// TIA Portal project "liftvezerles" (V17)
// Az Automatizálási Tanszék SIMATIC eszközei

(* hardware
DEVICE "S7-1200 station_1"  S7-1200 Station
   slot 0: "Rack_0"  S7-1200 Rack  Rack  V1.0
   slot 1: "S71214_sim"  CPU 1214C DC/DC/DC  6ES7 214-1AG40-0XB0  V4.0
   slot 3: "AQ 1x12BIT_1"  AQ1 signal board  6ES7 232-4HA30-0XB0  V1.0
DEVICE "KTP700.Basic"  KTP700 Basic PN
   slot 0: "KTP700.Basic"  KTP700 Basic PN  6AV2 123-2GB03-0AX0  17.0.0.0
   slot 1: "HMI_RT_1"  KTP700 Basic PN  6AV2 123-2GB03-0AX0  17.0.0.0
   slot 5: "KTP700.Basic.IE_CP_1"  PROFINET Interface  17.0.0.0
      slot 1: "PROFINET Interface_1"  PROFINET Interface
         slot 1: "Port_1"  Port
DEVICE "S7-1200 station_2"  S7-1200 Station
   slot 0: "Rack_0"  S7-1200 Rack  Rack  V1.0
   slot 1: "S7.1214_aut"  CPU 1214C DC/DC/DC  6ES7 214-1AG31-0XB0  V3.0
   slot 3: "AQ 1x12BIT_1"  AQ1 signal board  6ES7 232-4HA30-0XB0  V1.0
*)

// ===== PLC "S71214_sim"  CPU 1214C DC/DC/DC =====

VAR_GLOBAL   // PLC tag table "Default tag table"
   "System_Byte" AT %MB11 : Byte;
   "FirstScan" AT %M11.0 : Bool;
   "DiagStatusUpdate" AT %M11.1 : Bool;
   "AlwaysTRUE" AT %M11.2 : Bool;
   "AlwaysFALSE" AT %M11.3 : Bool;
   "Clock_Byte" AT %MB10 : Byte;
   "Clock_10Hz" AT %M10.0 : Bool;
   "Clock_5Hz" AT %M10.1 : Bool;
   "Clock_2.5Hz" AT %M10.2 : Bool;
   "Clock_2Hz" AT %M10.3 : Bool;
   "Clock_1.25Hz" AT %M10.4 : Bool;
   "Clock_1Hz" AT %M10.5 : Bool;
   "Clock_0.625Hz" AT %M10.6 : Bool;
   "Clock_0.5Hz" AT %M10.7 : Bool;
END_VAR

VAR_GLOBAL   // PLC tag table "Elevatorcontrol"
   "elevator1position" AT %MW28 : Int;
   "elevator2position" AT %MW26 : Int;
END_VAR

VAR_GLOBAL   // PLC tag table "IO"
   "door1closemotor" AT %M8.0 : Bool;
   "door2openmotor" AT %M8.1 : Bool;
   "door1opensens" AT %M8.2 : Bool;
   "door1closedsens" AT %M8.3 : Bool;
   "door2opensens" AT %M8.4 : Bool;
   "door2closedsens" AT %M8.5 : Bool;
   "door1openmotor" AT %M8.6 : Bool;
   "door2closemotor" AT %M8.7 : Bool;
   "elevator1upmotor" AT %M9.0 : Bool;
   "elevator1downmotor" AT %M9.1 : Bool;
   "elevator2upmotor" AT %M9.2 : Bool;
   "elevator2downmotor" AT %M9.3 : Bool;
   "proximity1ground" AT %M9.4 : Bool;
   "proximity11" AT %M9.5 : Bool;
   "proximity12" AT %M9.6 : Bool;
   "proximity13" AT %M9.7 : Bool;
   "proximity14" AT %M12.0 : Bool;
   "proximity15" AT %M12.1 : Bool;
   "proximity2ground" AT %M12.2 : Bool;
   "proximity21" AT %M12.3 : Bool;
   "proximity22" AT %M12.4 : Bool;
   "proximity23" AT %M12.5 : Bool;
   "proximity24" AT %M12.6 : Bool;
   "proximity25" AT %M12.7 : Bool;
END_VAR

VAR_GLOBAL   // PLC tag table "HMI_IO"
   "requpgnd" AT %M7.0 : Bool;
   "requp1" AT %M7.1 : Bool;
   "requp2" AT %M7.2 : Bool;
   "requp3" AT %M7.3 : Bool;
   "requp4" AT %M7.4 : Bool;
   "reqdown5" AT %M7.5 : Bool;
   "reqdown4" AT %M7.6 : Bool;
   "reqdown3" AT %M7.7 : Bool;
   "reqdown2" AT %M5.6 : Bool;
   "reqdown1" AT %M5.7 : Bool;
   "req10" AT %M4.2 : Bool;
   "req11" AT %M4.3 : Bool;
   "req12" AT %M4.4 : Bool;
   "req13" AT %M4.5 : Bool;
   "req14" AT %M4.6 : Bool;
   "req15" AT %M4.7 : Bool;
   "req20" AT %M5.0 : Bool;
   "req21" AT %M5.1 : Bool;
   "req22" AT %M5.2 : Bool;
   "req23" AT %M5.3 : Bool;
   "req24" AT %M5.4 : Bool;
   "req25" AT %M5.5 : Bool;
   "las2" AT %M6.1 : Bool;
   "las1" AT %M6.0 : Bool;
   "doorclosebutton1" AT %M6.2 : Bool;
   "doorclosebutton2" AT %M6.3 : Bool;
   "dooropenbutton1" AT %M6.4 : Bool;
   "dooropenbutton2" AT %M6.5 : Bool;
END_VAR

VAR_GLOBAL   // PLC tag table "IO_simulation_tags"
   "lastfloor1" AT %MW18 : Int;
   "lastfloor2" AT %MW20 : Int;
   "state1" AT %MW22 : Int;
   "state2" AT %MW24 : Int;
   "elevator1positionsim" AT %MW14 : Int;
   "elevator2positionsim" AT %MW16 : Int;
END_VAR

VAR_GLOBAL   // PLC tag table "HMI_display_tags"
   "activefloor" AT %MW40 : Int;
   "door1open" AT %M42.0 : Bool;
   "door2open" AT %M42.1 : Bool;
END_VAR

DATA_BLOCK "ControlBlock_DB"   // DB9
{ S7_Optimized_Access := 'TRUE' }
VERSION : 0.1
// stored: InstanceOfName ControlBlock
"ControlBlock"
BEGIN
END_DATA_BLOCK

// folder: System blocks/Program resources

DATA_BLOCK "door1closing"   // DB5
{ S7_Optimized_Access := 'TRUE' }
AUTHOR : Simatic
FAMILY : IEC
NAME : IEC_TMR
VERSION : 1.0
// stored: InstanceOfName IEC_TIMER
"IEC_TIMER"
BEGIN
END_DATA_BLOCK

DATA_BLOCK "door1opening"   // DB6
{ S7_Optimized_Access := 'TRUE' }
AUTHOR : Simatic
FAMILY : IEC
NAME : IEC_TMR
VERSION : 1.0
// stored: InstanceOfName IEC_TIMER
"IEC_TIMER"
BEGIN
END_DATA_BLOCK

DATA_BLOCK "door2closing"   // DB7
{ S7_Optimized_Access := 'TRUE' }
AUTHOR : Simatic
FAMILY : IEC
NAME : IEC_TMR
VERSION : 1.0
// stored: InstanceOfName IEC_TIMER
"IEC_TIMER"
BEGIN
END_DATA_BLOCK

DATA_BLOCK "door2opening"   // DB8
{ S7_Optimized_Access := 'TRUE' }
AUTHOR : Simatic
FAMILY : IEC
NAME : IEC_TMR
VERSION : 1.0
// stored: InstanceOfName IEC_TIMER
"IEC_TIMER"
BEGIN
END_DATA_BLOCK

DATA_BLOCK "starting_up2"   // DB10
{ S7_Optimized_Access := 'TRUE' }
AUTHOR : Simatic
FAMILY : IEC
NAME : IEC_TMR
VERSION : 1.0
// stored: InstanceOfName IEC_TIMER
"IEC_TIMER"
BEGIN
END_DATA_BLOCK

DATA_BLOCK "starting_down2"   // DB11
{ S7_Optimized_Access := 'TRUE' }
AUTHOR : Simatic
FAMILY : IEC
NAME : IEC_TMR
VERSION : 1.0
// stored: InstanceOfName IEC_TIMER
"IEC_TIMER"
BEGIN
END_DATA_BLOCK

DATA_BLOCK "goingup2"   // DB12
{ S7_Optimized_Access := 'TRUE' }
AUTHOR : Simatic
FAMILY : IEC
NAME : IEC_TMR
VERSION : 1.0
// stored: InstanceOfName IEC_TIMER
"IEC_TIMER"
BEGIN
END_DATA_BLOCK

DATA_BLOCK "goingdown2"   // DB13
{ S7_Optimized_Access := 'TRUE' }
AUTHOR : Simatic
FAMILY : IEC
NAME : IEC_TMR
VERSION : 1.0
// stored: InstanceOfName IEC_TIMER
"IEC_TIMER"
BEGIN
END_DATA_BLOCK

DATA_BLOCK "starting_up1"   // DB20
{ S7_Optimized_Access := 'TRUE' }
AUTHOR : Simatic
FAMILY : IEC
NAME : IEC_TMR
VERSION : 1.0
// stored: InstanceOfName IEC_TIMER
"IEC_TIMER"
BEGIN
END_DATA_BLOCK

DATA_BLOCK "starting_down1"   // DB21
{ S7_Optimized_Access := 'TRUE' }
AUTHOR : Simatic
FAMILY : IEC
NAME : IEC_TMR
VERSION : 1.0
// stored: InstanceOfName IEC_TIMER
"IEC_TIMER"
BEGIN
END_DATA_BLOCK

DATA_BLOCK "goingup1"   // DB22
{ S7_Optimized_Access := 'TRUE' }
AUTHOR : Simatic
FAMILY : IEC
NAME : IEC_TMR
VERSION : 1.0
// stored: InstanceOfName IEC_TIMER
"IEC_TIMER"
BEGIN
END_DATA_BLOCK

DATA_BLOCK "goingdown1"   // DB23
{ S7_Optimized_Access := 'TRUE' }
AUTHOR : Simatic
FAMILY : IEC
NAME : IEC_TMR
VERSION : 1.0
// stored: InstanceOfName IEC_TIMER
"IEC_TIMER"
BEGIN
END_DATA_BLOCK

// folder: (top level)

FUNCTION_BLOCK "Elevator"   // FB1, SCL
{ S7_Optimized_Access := 'TRUE' }
VERSION : 0.1
   VAR_INPUT
      doorclosedsens : Bool;
      dooropensens : Bool;
      currentlevel : Int := 5;
      nextlevel : Int := 0;
      las : Bool := true;
      closethedoorbutton : Bool;
      ack : Bool;
      stopidling : Bool;
      openthedoorbutton : Bool;
   END_VAR
   VAR_OUTPUT
      idling : Bool;
      opendoor : Bool;
      closedoor : Bool;
      headingup : Bool;
      headingdown : Bool;
      callcompleted : Bool;
   END_VAR
   VAR
      state : Int;
      idlewait : TON_TIME;
      closedoorwait : TON_TIME;
   END_VAR
BEGIN
   //states:
   //0: default
   //1: idle with doors closed
   //2: opening doors
   //3: opendoors, waiting to close
   //4: closing doors
   //5: going down
   //6: going up
   //7: arrived, opening door
   //8: arrived, door opened
   //20: idling with doors opened
   //21: idling, closing doors


   #idlewait(IN:=(#state = 20 AND #las),
             PT:=T#20s);
   #closedoorwait(IN:=((#state = 3) AND #las),
                  PT:=T#5s);




   CASE #state OF
       0:
           IF #currentlevel = 0 AND #doorclosedsens THEN
               #state := 21;
           END_IF;
       1:
           IF NOT(#currentlevel = #nextlevel) THEN
               #state := 3;
           END_IF;
       2:
           IF #dooropensens THEN
               #state := 3;
           END_IF;


       3:
           IF #closedoorwait.Q OR #closethedoorbutton THEN
               #state := 4;
           END_IF;
       4:
           IF #doorclosedsens AND #currentlevel>#nextlevel THEN
               #state := 5;
           ELSIF #doorclosedsens AND #currentlevel<#nextlevel THEN
               #state := 6;
           ELSIF #doorclosedsens AND #currentlevel=#nextlevel THEN
               #state := 7;
           ELSIF NOT #las THEN
               #state := 3;
           END_IF;
       5,6:
           IF #currentlevel=#nextlevel THEN
               #state := 7;
           END_IF;
       7:
           IF #dooropensens THEN
               #state := 8;
           END_IF;
       8: IF #ack THEN
               #callcompleted := FALSE;
               #state := 20;
               END_IF;
           #callcompleted := TRUE;


       20:
           IF NOT(#currentlevel = #nextlevel) THEN
               #state := 3;
           ELSIF (#idlewait.Q OR #closethedoorbutton) THEN
               #state := 21;
           END_IF;
       21:
           IF #stopidling THEN
               #state := 7;
           ELSIF NOT(#currentlevel = #nextlevel) THEN
               IF #doorclosedsens AND #currentlevel > #nextlevel THEN
                   #state := 5;
               ELSIF #doorclosedsens AND #currentlevel < #nextlevel THEN
                   #state := 6;
               END_IF;
           ELSIF #openthedoorbutton THEN
               #state := 20;
           END_IF;
       ELSE
           #state := 0;

   END_CASE;

   #callcompleted := (#state = 8 OR #state=3);
   #headingup := (#state = 6);
   #headingdown := (#state = 5) OR (#state = 0);
   #closedoor := (#state = 4) OR (#state = 21) OR (#state=0) OR (#state=1) OR (#state=5) OR (#state=6);
   #opendoor := (#state = 2) OR (#state = 7) OR (#state=3) OR (#state=20) OR (#state=8);
   #idling := #state = 21;
END_FUNCTION_BLOCK

FUNCTION_BLOCK "ControlBlock"   // FB2, SCL
{ S7_Optimized_Access := 'TRUE' }
VERSION : 0.1
   VAR
      requparray : Array[0..5] of Bool;
      reqdownarray : Array[0..5] of Bool;
      elevator1reqarray : Array[0..5] of Bool;
      elevator2reqarray : Array[0..5] of Bool;
      elevator1next : Int := 0;
      elevator2next : Int := 0;
      elevator1heading : Int;
      elevator2heading : Int;
      elevator1 : "Elevator";
      elevator2 : "Elevator";
      elevator1ack : Bool;
      elevator2ack : Bool;
      elevator1stopidling : Bool;
      elevator2stopidling : Bool;
      elevator1distance : Int;
      elevator2distance : Int;
      reqlocation : Int;
   END_VAR
BEGIN
   // "sensors_to_int_position"(in1g:="proximity1ground",
   //                           in11:="proximity11",
   //                           in12:="proximity12",
   //                           in13:="proximity13",
   //                           in14:="proximity14",
   //                           in15:="proximity15",
   //                           in2g:="proximity2ground",
   //                           in21:="proximity21",
   //                           in22:="proximity22",
   //                           in23:="proximity23",
   //                           in24:="proximity24",
   //                           in25:="proximity25",
   //                           out1=>"elevator1position",
   //                           out2=>"elevator2position");

   IF "proximity1ground" THEN
       "elevator1position" := 0;
   END_IF;
   IF "proximity11" THEN
       "elevator1position" := 1;
   END_IF;
   IF "proximity12" THEN
       "elevator1position" := 2;
   END_IF;
   IF "proximity13" THEN
       "elevator1position" := 3;
   END_IF;
   IF "proximity14" THEN
       "elevator1position" := 4;
   END_IF;
   IF "proximity15" THEN
       "elevator1position" := 5;
   END_IF;

   IF "proximity2ground" THEN
       "elevator2position" := 0;
   END_IF;
   IF "proximity21" THEN
       "elevator2position" := 1;
   END_IF;
   IF "proximity22" THEN
       "elevator2position" := 2;
   END_IF;
   IF "proximity23" THEN
       "elevator2position" := 3;
   END_IF;
   IF "proximity24" THEN
       "elevator2position" := 4;
   END_IF;
   IF "proximity25" THEN
       "elevator2position" := 5;
   END_IF;




   //heading:
   //0: idle
   //1: down
   //2: up


   IF #elevator1.callcompleted THEN
       CASE "elevator1position" OF
           0:
               "req10" := FALSE;
               "requpgnd" := FALSE;
           1:
               "req11" := FALSE;
               "requp1" := FALSE;
               "reqdown1" := FALSE;
           2:
               "req12" := FALSE;
               "requp2" := FALSE;
               "reqdown2" := FALSE;
           3:
               "req13" := FALSE;
               "requp3" := FALSE;
               "reqdown3" := FALSE;
           4:
               "req14" := FALSE;
               "requp4" := FALSE;
               "reqdown4" := FALSE;
           5:
               "req15" := FALSE;
               "reqdown5" := FALSE;
       END_CASE;
       #elevator1ack := TRUE;
   ELSE
       #elevator1ack := FALSE;
   END_IF;


   IF #elevator2.callcompleted THEN
       CASE "elevator2position" OF
           0:
               "req20" := FALSE;
               "requpgnd" := FALSE;
           1:
               "req21" := FALSE;
               "requp1" := FALSE;
               "reqdown1" := FALSE;
           2:
               "req22" := FALSE;
               "requp2" := FALSE;
               "reqdown2" := FALSE;
           3:
               "req23" := FALSE;
               "requp3" := FALSE;
               "reqdown3" := FALSE;
           4:
               "req24" := FALSE;
               "requp4" := FALSE;
               "reqdown4" := FALSE;
           5:
               "req25" := FALSE;
               "reqdown5" := FALSE;

       END_CASE;

       #elevator2ack := TRUE;
   ELSE
       #elevator2ack := FALSE;
   END_IF;
   // distance calculation, if both idle:
   IF ((#elevator1heading = 0 AND #elevator2heading = 0) AND ("requpgnd" OR "requp2" OR "requp3" OR "requp4" OR "reqdown5" OR "reqdown4" OR "reqdown3" OR "reqdown2" OR "reqdown1")) THEN
       IF "requpgnd" THEN
           #elevator1distance := "elevator1position";
           #elevator2distance := "elevator2position";
           #reqlocation := 0;
           "requpgnd" := FALSE;
       END_IF;
       IF ("requp1" OR "reqdown1") THEN
           #elevator1distance := ABS("elevator1position" - 1);
           #elevator2distance := ABS("elevator2position" - 1);
           #reqlocation := 1;
           "requp1" := FALSE;
           "reqdown1" := FALSE;
       END_IF;
       IF ("requp2" OR "reqdown2") THEN
           #elevator1distance := ABS("elevator1position" - 2);
           #elevator2distance := ABS("elevator2position" - 2);
           #reqlocation := 2;
           "requp2" := FALSE;
           "reqdown2" := FALSE;
       END_IF;
       IF ("requp3" OR "reqdown3") THEN
           #elevator1distance := ABS("elevator1position" - 3);
           #elevator2distance := ABS("elevator2position" - 3);
           #reqlocation := 3;
           "requp3" := FALSE;
           "reqdown3" := FALSE;
       END_IF;
       IF ("requp4" OR "reqdown4") THEN
           #elevator1distance := ABS("elevator1position" - 4);
           #elevator2distance := ABS("elevator2position" - 4);
           #reqlocation := 4;
           "requp4" := FALSE;
           "reqdown4" := FALSE;
       END_IF;
       IF "reqdown5" THEN
           #elevator1distance := 5 - "elevator1position";
           #elevator2distance := 5 - "elevator2position";
           #reqlocation := 5;
           "reqdown5" := FALSE;
       END_IF;

       IF (#elevator1distance > #elevator2distance) THEN
           #elevator2next := #reqlocation;
           CASE #reqlocation OF
               0:
                   "req20" := TRUE;
               1:
                   "req21" := TRUE;
               2:
                   "req22" := TRUE;
               3:
                   "req23" := TRUE;
               4:
                   "req24" := TRUE;
               5:
                   "req25" := TRUE;

           END_CASE;


       ELSE
           #elevator1next := #reqlocation;
           CASE #reqlocation OF
               0:
                   "req10" := TRUE;
               1:
                   "req11" := TRUE;
               2:
                   "req12" := TRUE;
               3:
                   "req13" := TRUE;
               4:
                   "req14" := TRUE;
               5:
                   "req15" := TRUE;

           END_CASE;

       END_IF;

       ;

       ELSE
       //ELEVATOR1:


       IF (#elevator1heading = 2) OR (#elevator1heading = 0) THEN             //felfelé lift 1
           CASE "elevator1position" OF
               0:
                   IF (("req10" OR "requpgnd") AND "proximity1ground") THEN
                       #elevator1next := 0;
                   ELSIF ("req11" OR "requp1") THEN
                       #elevator1next := 1;
                       #elevator1heading := 2;
                   ELSIF ("req12" OR "requp2") THEN
                       #elevator1next := 2;
                       #elevator1heading := 2;
                   ELSIF ("req13" OR "requp3") THEN
                       #elevator1next := 3;
                       #elevator1heading := 2;
                   ELSIF ("req14" OR "requp4") THEN
                       #elevator1next := 4;
                       #elevator1heading := 2;
                   ELSIF ("req15") THEN
                       #elevator1next := 5;
                       #elevator1heading := 2;
                   ELSIF ("reqdown5") THEN
                       "reqdown5" := FALSE;
                       "req15" := TRUE;
                       #elevator1next := 5;
                       #elevator1heading := 2;
                   ELSIF ("reqdown4") THEN
                       "reqdown4" := FALSE;
                       "req14" := TRUE;
                       #elevator1next := 4;
                       #elevator1heading := 2;
                   ELSIF ("reqdown3") THEN
                       "reqdown3" := FALSE;
                       "req13" := TRUE;
                       #elevator1next := 3;
                       #elevator1heading := 2;
                   ELSIF ("reqdown2") THEN
                       "reqdown4" := FALSE;
                       "req12" := TRUE;
                       #elevator1next := 2;
                       #elevator1heading := 2;
                   ELSIF ("reqdown1") THEN
                       "reqdown1" := FALSE;
                       "req11" := TRUE;
                       #elevator1next := 1;
                       #elevator1heading := 2;
                   ELSE
                       #elevator1heading := 0;
                   END_IF;

               1:
                   IF (("req11" OR "requp1") AND "proximity11") THEN
                       #elevator1next := 1;
                   ELSIF ("req12" OR "requp2") THEN
                       #elevator1next := 2;
                       #elevator1heading := 2;
                   ELSIF ("req13" OR "requp3") THEN
                       #elevator1next := 3;
                       #elevator1heading := 2;
                   ELSIF ("req14" OR "requp4") THEN
                       #elevator1next := 4;
                       #elevator1heading := 2;
                   ELSIF ("req15") THEN
                       #elevator1next := 5;
                       #elevator1heading := 2;
                   ELSIF ("reqdown5") THEN
                       "reqdown5" := FALSE;
                       "req15" := TRUE;
                       #elevator1next := 5;
                       #elevator1heading := 2;
                   ELSIF ("reqdown4") THEN
                       "reqdown4" := FALSE;
                       "req14" := TRUE;
                       #elevator1next := 4;
                       #elevator1heading := 2;
                   ELSIF ("reqdown3") THEN
                       "reqdown3" := FALSE;
                       "req13" := TRUE;
                       #elevator1next := 3;
                       #elevator1heading := 2;
                   ELSIF ("reqdown2") THEN
                       "reqdown4" := FALSE;
                       "req12" := TRUE;
                       #elevator1next := 2;
                       #elevator1heading := 2;
                   ELSE
                       #elevator1heading := 0;
                   END_IF;

               2:
                   IF (("req12" OR "requp2") AND "proximity12") THEN
                       #elevator1next := 2;
                   ELSIF ("req13" OR "requp3") THEN
                       #elevator1next := 3;
                       #elevator1heading := 2;
                   ELSIF ("req14" OR "requp4") THEN
                       #elevator1next := 4;
                       #elevator1heading := 2;
                   ELSIF ("req15") THEN
                       #elevator1next := 5;
                       #elevator1heading := 2;
                   ELSIF ("reqdown5") THEN
                       "reqdown5" := FALSE;
                       "req15" := TRUE;
                       #elevator1next := 5;
                       #elevator1heading := 2;
                   ELSIF ("reqdown4") THEN
                       "reqdown4" := FALSE;
                       "req14" := TRUE;
                       #elevator1next := 4;
                       #elevator1heading := 2;
                   ELSIF ("reqdown3") THEN
                       "reqdown3" := FALSE;
                       "req13" := TRUE;
                       #elevator1next := 3;
                       #elevator1heading := 2;
                   ELSE
                       #elevator1heading := 0;
                   END_IF;

               3:
                   IF (("req13" OR "requp3" AND "proximity13")) THEN
                       #elevator1next := 3;
                   ELSIF ("req14" OR "requp4") THEN
                       #elevator1next := 4;
                       #elevator1heading := 2;
                   ELSIF ("req15") THEN
                       #elevator1next := 5;
                       #elevator1heading := 2;
                   ELSIF ("reqdown5") THEN
                       "reqdown5" := FALSE;
                       "req15" := TRUE;
                       #elevator1next := 5;
                       #elevator1heading := 2;
                   ELSIF ("reqdown4") THEN
                       "reqdown4" := FALSE;
                       "req14" := TRUE;
                       #elevator1next := 4;
                       #elevator1heading := 2;
                   ELSE
                       #elevator1heading := 0;
                   END_IF;
                   ;
               4:
                   IF (("req14" OR "requp4") AND "proximity14") THEN
                       #elevator1next := 4;
                   ELSIF ("req15") THEN
                       #elevator1next := 5;
                       #elevator1heading := 2;
                   ELSIF ("reqdown5") THEN
                       "reqdown5" := FALSE;
                       "req15" := TRUE;
                       #elevator1next := 5;
                       #elevator1heading := 2;
                   ELSE
                       #elevator1heading := 0;
                   END_IF;

               5:
                   IF ("req15" AND "proximity15") THEN
                       #elevator1next := 5;
                   END_IF;
                   #elevator1heading := 0;
           END_CASE;

           ;
       END_IF;


       IF (#elevator1heading = 1) OR (#elevator1heading = 0) THEN             //lefelé lift1
           CASE "elevator1position" OF
               0:
                   IF ("req10" AND "proximity1ground") THEN
                       #elevator1next := 0;
                   END_IF;
                   #elevator1heading := 0;

               1:
                   IF (("req11" OR "reqdown1") AND "proximity11") THEN
                       #elevator1next := 1;
                   ELSIF ("req10") THEN
                       #elevator1next := 0;
                       #elevator1heading := 1;
                   ELSIF ("requpgnd") THEN
                       "requpgnd" := FALSE;
                       "req10" := TRUE;
                       #elevator1next := 0;
                       #elevator1heading := 1;
                   ELSE
                       #elevator1heading := 0;
                   END_IF;

               2:
                   IF (("req12" OR "reqdown2") AND "proximity12") THEN
                       #elevator1next := 2;
                   ELSIF ("req11" OR "reqdown1") THEN
                       #elevator1next := 1;
                       #elevator1heading := 1;
                   ELSIF ("req10") THEN
                       #elevator1next := 0;
                       #elevator1heading := 1;
                   ELSIF ("requpgnd") THEN
                       "requpgnd" := FALSE;
                       "req10" := TRUE;
                       #elevator1next := 0;
                       #elevator1heading := 1;
                   ELSIF ("requp1") THEN
                       "requp1" := FALSE;
                       "req11" := TRUE;
                       #elevator1next := 1;
                       #elevator1heading := 1;
                   ELSE
                       #elevator1heading := 0;
                   END_IF;

               3:
                   IF (("req13" OR "reqdown3") AND "proximity13") THEN
                       #elevator1next := 3;
                   ELSIF ("req12" OR "reqdown2") THEN
                       #elevator1next := 2;
                       #elevator1heading := 1;
                   ELSIF ("req11" OR "reqdown1") THEN
                       #elevator1next := 1;
                       #elevator1heading := 1;
                   ELSIF ("req10") THEN
                       #elevator1next := 0;
                       #elevator1heading := 1;
                   ELSIF ("requpgnd") THEN
                       "requpgnd" := FALSE;
                       "req10" := TRUE;
                       #elevator1next := 0;
                       #elevator1heading := 1;
                   ELSIF ("requp1") THEN
                       "requp1" := FALSE;
                       "req11" := TRUE;
                       #elevator1next := 1;
                       #elevator1heading := 1;
                   ELSIF ("requp2") THEN
                       "requp2" := FALSE;
                       "req12" := TRUE;
                       #elevator1next := 2;
                       #elevator1heading := 1;
                   ELSE
                       #elevator1heading := 0;
                   END_IF;
               4:
                   IF (("req14" OR "reqdown4") AND "proximity14") THEN
                       #elevator1next := 4;
                   ELSIF ("req13" OR "reqdown3") THEN
                       #elevator1next := 3;
                       #elevator1heading := 1;
                   ELSIF ("req12" OR "reqdown2") THEN
                       #elevator1next := 2;
                       #elevator1heading := 1;
                   ELSIF ("req11" OR "reqdown1") THEN
                       #elevator1next := 1;
                       #elevator1heading := 1;
                   ELSIF ("req10") THEN
                       #elevator1next := 0;
                       #elevator1heading := 1;
                   ELSIF ("requpgnd") THEN
                       "requpgnd" := FALSE;
                       "req10" := TRUE;
                       #elevator1next := 0;
                       #elevator1heading := 1;
                   ELSIF ("requp1") THEN
                       "requp1" := FALSE;
                       "req11" := TRUE;
                       #elevator1next := 1;
                       #elevator1heading := 1;
                   ELSIF ("requp2") THEN
                       "requp2" := FALSE;
                       "req12" := TRUE;
                       #elevator1next := 2;
                       #elevator1heading := 1;
                   ELSIF ("requp3") THEN
                       "requp3" := FALSE;
                       "req13" := TRUE;
                       #elevator1next := 3;
                       #elevator1heading := 1;
                   ELSE
                       #elevator1heading := 0;
                   END_IF;

               5:
                   IF (("req15" OR "reqdown5") AND "proximity15") THEN
                       #elevator1next := 5;
                   ELSIF ("req14" OR "reqdown4") THEN
                       #elevator1next := 4;
                       #elevator1heading := 1;
                   ELSIF ("req13" OR "reqdown3") THEN
                       #elevator1next := 3;
                       #elevator1heading := 1;
                   ELSIF ("req12" OR "reqdown2") THEN
                       #elevator1next := 2;
                       #elevator1heading := 1;
                   ELSIF ("req11" OR "reqdown1") THEN
                       #elevator1next := 1;
                       #elevator1heading := 1;
                   ELSIF ("req10") THEN
                       #elevator1next := 0;
                       #elevator1heading := 1;
                   ELSIF ("requpgnd") THEN
                       "requpgnd" := FALSE;
                       "req10" := TRUE;
                       #elevator1next := 0;
                       #elevator1heading := 1;
                   ELSIF ("requp1") THEN
                       "requp1" := FALSE;
                       "req11" := TRUE;
                       #elevator1next := 1;
                       #elevator1heading := 1;
                   ELSIF ("requp2") THEN
                       "requp2" := FALSE;
                       "req12" := TRUE;
                       #elevator1next := 2;
                       #elevator1heading := 1;
                   ELSIF ("requp3") THEN
                       "requp3" := FALSE;
                       "req13" := TRUE;
                       #elevator1next := 3;
                       #elevator1heading := 1;
                   ELSIF ("requp4") THEN
                       "requp4" := FALSE;
                       "req14" := TRUE;
                       #elevator1next := 4;
                       #elevator1heading := 1;

                   ELSE
                       #elevator1heading := 0;
                   END_IF;
           END_CASE;

           ;
       END_IF;

       //"Elevator2"


       IF (#elevator2heading = 2) OR (#elevator2heading = 0) THEN             //felfelé lift 2
           CASE "elevator2position" OF
               0:
                   IF (("req20" OR "requpgnd") AND "proximity2ground") THEN
                       #elevator2next := 0;
                   ELSIF ("req21" OR "requp1") THEN
                       #elevator2next := 1;
                       #elevator2heading := 2;
                   ELSIF ("req22" OR "requp2") THEN
                       #elevator2next := 2;
                       #elevator2heading := 2;
                   ELSIF ("req23" OR "requp3") THEN
                       #elevator2next := 3;
                       #elevator2heading := 2;
                   ELSIF ("req24" OR "requp4") THEN
                       #elevator2next := 4;
                       #elevator2heading := 2;
                   ELSIF ("req25") THEN
                       #elevator2next := 5;
                       #elevator2heading := 2;
                   ELSIF ("reqdown5") THEN
                       "reqdown5" := FALSE;
                       "req25" := TRUE;
                       #elevator2next := 5;
                       #elevator2heading := 2;
                   ELSIF ("reqdown4") THEN
                       "reqdown4" := FALSE;
                       "req24" := TRUE;
                       #elevator2next := 4;
                       #elevator2heading := 2;
                   ELSIF ("reqdown3") THEN
                       "reqdown3" := FALSE;
                       "req23" := TRUE;
                       #elevator2next := 3;
                       #elevator2heading := 2;
                   ELSIF ("reqdown2") THEN
                       "reqdown4" := FALSE;
                       "req22" := TRUE;
                       #elevator2next := 2;
                       #elevator2heading := 2;
                   ELSIF ("reqdown1") THEN
                       "reqdown1" := FALSE;
                       "req21" := TRUE;
                       #elevator2next := 1;
                       #elevator2heading := 2;
                   ELSE
                       #elevator2heading := 0;
                   END_IF;

               1:
                   IF (("req21" OR "requp1") AND "proximity21") THEN
                       #elevator2next := 1;
                   ELSIF ("req22" OR "requp2") THEN
                       #elevator2next := 2;
                       #elevator2heading := 2;
                   ELSIF ("req23" OR "requp3") THEN
                       #elevator2next := 3;
                       #elevator2heading := 2;
                   ELSIF ("req24" OR "requp4") THEN
                       #elevator2next := 4;
                       #elevator2heading := 2;
                   ELSIF ("req25") THEN
                       #elevator2next := 5;
                       #elevator2heading := 2;
                   ELSIF ("reqdown5") THEN
                       "reqdown5" := FALSE;
                       "req25" := TRUE;
                       #elevator2next := 5;
                       #elevator2heading := 2;
                   ELSIF ("reqdown4") THEN
                       "reqdown4" := FALSE;
                       "req24" := TRUE;
                       #elevator2next := 4;
                       #elevator2heading := 2;
                   ELSIF ("reqdown3") THEN
                       "reqdown3" := FALSE;
                       "req23" := TRUE;
                       #elevator2next := 3;
                       #elevator2heading := 2;
                   ELSIF ("reqdown2") THEN
                       "reqdown4" := FALSE;
                       "req22" := TRUE;
                       #elevator2next := 2;
                       #elevator2heading := 2;
                   ELSE
                       #elevator2heading := 0;
                   END_IF;

               2:
                   IF (("req22" OR "requp2") AND "proximity22") THEN
                       #elevator2next := 2;
                   ELSIF ("req23" OR "requp3") THEN
                       #elevator2next := 3;
                       #elevator2heading := 2;
                   ELSIF ("req24" OR "requp4") THEN
                       #elevator2next := 4;
                       #elevator2heading := 2;
                   ELSIF ("req25") THEN
                       #elevator2next := 5;
                       #elevator2heading := 2;
                   ELSIF ("reqdown5") THEN
                       "reqdown5" := FALSE;
                       "req25" := TRUE;
                       #elevator2next := 5;
                       #elevator2heading := 2;
                   ELSIF ("reqdown4") THEN
                       "reqdown4" := FALSE;
                       "req24" := TRUE;
                       #elevator2next := 4;
                       #elevator2heading := 2;
                   ELSIF ("reqdown3") THEN
                       "reqdown3" := FALSE;
                       "req23" := TRUE;
                       #elevator2next := 3;
                       #elevator2heading := 2;
                   ELSE
                       #elevator2heading := 0;
                   END_IF;

               3:
                   IF (("req23" OR "requp3") AND "proximity23") THEN
                       #elevator2next := 3;
                   ELSIF ("req24" OR "requp4") THEN
                       #elevator2next := 4;
                       #elevator2heading := 2;
                   ELSIF ("req25") THEN
                       #elevator2next := 5;
                       #elevator2heading := 2;
                   ELSIF ("reqdown5") THEN
                       "reqdown5" := FALSE;
                       "req25" := TRUE;
                       #elevator2next := 5;
                       #elevator2heading := 2;
                   ELSIF ("reqdown4") THEN
                       "reqdown4" := FALSE;
                       "req24" := TRUE;
                       #elevator2next := 4;
                       #elevator2heading := 2;
                   ELSE
                       #elevator2heading := 0;
                   END_IF;
                   ;
               4:
                   IF (("req24" OR "requp4") AND "proximity24") THEN
                       #elevator2next := 4;
                   ELSIF ("req25") THEN
                       #elevator2next := 5;
                       #elevator2heading := 2;
                   ELSIF ("reqdown5") THEN
                       "reqdown5" := FALSE;
                       "req25" := TRUE;
                       #elevator2next := 5;
                       #elevator2heading := 2;
                   ELSE
                       #elevator2heading := 0;
                   END_IF;

               5:
                   IF ("req25" AND "proximity25") THEN
                       #elevator2next := 5;
                   END_IF;
                   #elevator2heading := 0;
           END_CASE;

           ;
       END_IF;


       IF (#elevator2heading = 1) OR (#elevator2heading = 0) THEN             //lefelé lift 2
           CASE "elevator2position" OF
               0:
                   IF ("req20" AND "proximity2ground") THEN
                       #elevator2next := 0;
                   END_IF;
                   #elevator2heading := 0;

               1:
                   IF (("req21" OR "reqdown1") AND "proximity21") THEN
                       #elevator2next := 1;
                   ELSIF ("req20") THEN
                       #elevator2next := 0;
                       #elevator2heading := 1;
                   ELSIF ("requpgnd") THEN
                       "requpgnd" := FALSE;
                       "req20" := TRUE;
                       #elevator2next := 0;
                       #elevator2heading := 1;
                   ELSE
                       #elevator2heading := 0;
                   END_IF;

               2:
                   IF (("req22" OR "reqdown2") AND "proximity22") THEN
                       #elevator2next := 2;
                   ELSIF ("req21" OR "reqdown1") THEN
                       #elevator2next := 1;
                       #elevator2heading := 1;
                   ELSIF ("req20") THEN
                       #elevator2next := 0;
                       #elevator2heading := 1;
                   ELSIF ("requpgnd") THEN
                       "requpgnd" := FALSE;
                       "req20" := TRUE;
                       #elevator2next := 0;
                       #elevator2heading := 1;
                   ELSIF ("requp1") THEN
                       "requp1" := FALSE;
                       "req21" := TRUE;
                       #elevator2next := 1;
                       #elevator2heading := 1;
                   ELSE
                       #elevator2heading := 0;
                   END_IF;

               3:
                   IF (("req23" OR "reqdown3") AND "proximity23") THEN
                       #elevator2next := 3;
                   ELSIF ("req22" OR "reqdown2") THEN
                       #elevator2next := 2;
                       #elevator2heading := 1;
                   ELSIF ("req21" OR "reqdown1") THEN
                       #elevator2next := 1;
                       #elevator2heading := 1;
                   ELSIF ("req20") THEN
                       #elevator2next := 0;
                       #elevator2heading := 1;
                   ELSIF ("requpgnd") THEN
                       "requpgnd" := FALSE;
                       "req20" := TRUE;
                       #elevator2next := 0;
                       #elevator2heading := 1;
                   ELSIF ("requp1") THEN
                       "requp1" := FALSE;
                       "req21" := TRUE;
                       #elevator2next := 1;
                       #elevator2heading := 1;
                   ELSIF ("requp2") THEN
                       "requp2" := FALSE;
                       "req22" := TRUE;
                       #elevator2next := 2;
                       #elevator2heading := 1;
                   ELSE
                       #elevator2heading := 0;
                   END_IF;
               4:
                   IF (("req24" OR "reqdown4") AND "proximity24") THEN
                       #elevator2next := 4;
                   ELSIF ("req23" OR "reqdown3") THEN
                       #elevator2next := 3;
                       #elevator2heading := 1;
                   ELSIF ("req22" OR "reqdown2") THEN
                       #elevator2next := 2;
                       #elevator2heading := 1;
                   ELSIF ("req21" OR "reqdown1") THEN
                       #elevator2next := 1;
                       #elevator2heading := 1;
                   ELSIF ("req20") THEN
                       #elevator2next := 0;
                       #elevator2heading := 1;
                   ELSIF ("requpgnd") THEN
                       "requpgnd" := FALSE;
                       "req20" := TRUE;
                       #elevator2next := 0;
                       #elevator2heading := 1;
                   ELSIF ("requp1") THEN
                       "requp1" := FALSE;
                       "req21" := TRUE;
                       #elevator2next := 1;
                       #elevator2heading := 1;
                   ELSIF ("requp2") THEN
                       "requp2" := FALSE;
                       "req22" := TRUE;
                       #elevator2next := 2;
                       #elevator2heading := 1;
                   ELSIF ("requp3") THEN
                       "requp3" := FALSE;
                       "req23" := TRUE;
                       #elevator2next := 3;
                       #elevator2heading := 1;
                   ELSE
                       #elevator2heading := 0;
                   END_IF;

               5:
                   IF (("req25" OR "reqdown5") AND "proximity25") THEN
                       #elevator2next := 5;
                   ELSIF ("req24" OR "reqdown4") THEN
                       #elevator2next := 4;
                       #elevator2heading := 1;
                   ELSIF ("req23" OR "reqdown3") THEN
                       #elevator2next := 3;
                       #elevator2heading := 1;
                   ELSIF ("req22" OR "reqdown2") THEN
                       #elevator2next := 2;
                       #elevator2heading := 1;
                   ELSIF ("req21" OR "reqdown1") THEN
                       #elevator2next := 1;
                       #elevator2heading := 1;
                   ELSIF ("req20") THEN
                       #elevator2next := 0;
                       #elevator2heading := 1;
                   ELSIF ("requpgnd") THEN
                       "requpgnd" := FALSE;
                       "req20" := TRUE;
                       #elevator2next := 0;
                       #elevator2heading := 1;
                   ELSIF ("requp1") THEN
                       "requp1" := FALSE;
                       "req21" := TRUE;
                       #elevator2next := 1;
                       #elevator2heading := 1;
                   ELSIF ("requp2") THEN
                       "requp2" := FALSE;
                       "req22" := TRUE;
                       #elevator2next := 2;
                       #elevator2heading := 1;
                   ELSIF ("requp3") THEN
                       "requp3" := FALSE;
                       "req23" := TRUE;
                       #elevator2next := 3;
                       #elevator2heading := 1;
                   ELSIF ("requp4") THEN
                       "requp4" := FALSE;
                       "req24" := TRUE;
                       #elevator2next := 4;
                       #elevator2heading := 1;

                   ELSE
                       #elevator2heading := 0;
                   END_IF;
           END_CASE;

           ;
       END_IF;

   END_IF;






       IF #elevator1.idling THEN
           CASE "elevator1position" OF
               0:
                   IF ("requpgnd" OR "req10") THEN
                       #elevator1stopidling := TRUE;
                   ELSE
                       #elevator1stopidling := FALSE;
                   END_IF;
                   ;
               1:
                   IF ("requp1" OR "reqdown1" OR "req11") THEN
                       #elevator1stopidling := TRUE;
                   ELSE
                       #elevator1stopidling := FALSE;
                   END_IF;
                   ;
               2:
                   IF ("requp2" OR "reqdown2" OR "req12") THEN
                       #elevator1stopidling := TRUE;
                   ELSE
                       #elevator1stopidling := FALSE;
                   END_IF;
                   ;
               3:
                   IF ("requp3" OR "reqdown3" OR "req13") THEN
                       #elevator1stopidling := TRUE;
                   ELSE
                       #elevator1stopidling := FALSE;
                   END_IF;
                   ;
               4:
                   IF ("requp4" OR "reqdown4" OR "req14") THEN
                       #elevator1stopidling := TRUE;
                   ELSE
                       #elevator1stopidling := FALSE;
                   END_IF;
                   ;
               5:
                   IF ("reqdown5" OR "req15") THEN
                       #elevator1stopidling := TRUE;
                   ELSE
                       #elevator1stopidling := FALSE;
                   END_IF;
                   ;
           END_CASE;

       END_IF;

       IF #elevator2.idling THEN
           CASE "elevator2position" OF
               0:
                   IF ("requpgnd" OR "req20") THEN
                       #elevator2stopidling := TRUE;
                   ELSE
                       #elevator2stopidling := FALSE;
                   END_IF;
                   ;
               1:
                   IF ("requp1" OR "reqdown1" OR "req21") THEN
                       #elevator2stopidling := TRUE;
                   ELSE
                       #elevator2stopidling := FALSE;
                   END_IF;
                   ;
               2:
                   IF ("requp2" OR "reqdown2" OR "req22") THEN
                       #elevator2stopidling := TRUE;
                   ELSE
                       #elevator2stopidling := FALSE;
                   END_IF;
                   ;
               3:
                   IF ("requp3" OR "reqdown3" OR "req23") THEN
                       #elevator2stopidling := TRUE;
                   ELSE
                       #elevator2stopidling := FALSE;
                   END_IF;
                   ;
               4:
                   IF ("requp4" OR "reqdown4" OR "req24") THEN
                       #elevator2stopidling := TRUE;
                   ELSE
                       #elevator2stopidling := FALSE;
                   END_IF;
                   ;
               5:
                   IF ("reqdown5" OR "req25") THEN
                       #elevator2stopidling := TRUE;
                   ELSE
                       #elevator2stopidling := FALSE;
                   END_IF;
                   ;
           END_CASE;

       END_IF;

   #elevator1(currentlevel:="elevator1position",
              doorclosedsens:="door1closedsens",
              dooropensens:="door1opensens",
              nextlevel:=#elevator1next,
              las:=true,
              stopidling:=#elevator1stopidling,
              closethedoorbutton:="doorclosebutton1",
              openthedoorbutton:="dooropenbutton1",
              ack:=#elevator1ack,
              opendoor=>"door1openmotor",
              closedoor=>"door1closemotor",
              headingup=>"elevator1upmotor",
              headingdown=>"elevator1downmotor");
   #elevator2(currentlevel:="elevator2position",
              doorclosedsens:="door2closedsens",
              dooropensens:="door2opensens",
              nextlevel:=#elevator2next,
              las:=TRUE,
              stopidling:=#elevator2stopidling,
              closethedoorbutton:="doorclosebutton2",
              openthedoorbutton:="dooropenbutton2",
              ack:=#elevator2ack,
              opendoor=>"door2openmotor",
              closedoor=>"door2closemotor",
              headingup=>"elevator2upmotor",
              headingdown=>"elevator2downmotor");
END_FUNCTION_BLOCK

FUNCTION "sensors_to_int_position" : Void   // FC1, SCL
{ S7_Optimized_Access := 'TRUE' }
VERSION : 0.1
   VAR_INPUT
      in1g : Bool;
      in11 : Bool;
      in12 : Bool;
      in13 : Bool;
      in14 : Bool;
      in15 : Bool;
      in2g : Bool;
      in21 : Bool;
      in22 : Bool;
      in23 : Bool;
      in24 : Bool;
      in25 : Bool;
   END_VAR
   VAR_OUTPUT
      out1 : Int;
      out2 : Int;
   END_VAR
BEGIN
   IF #in1g THEN
       #out1 := 0;
   END_IF;
   IF #in11 THEN
       #out1 := 1;
   END_IF;
   IF #in12 THEN
       #out1 := 2;
   END_IF;
   IF #in13 THEN
       #out1 := 3;
   END_IF;
   IF #in14 THEN
       #out1 := 4;
   END_IF;
   IF #in15 THEN
       #out1 := 5;
   END_IF;

   IF #in2g THEN
       #out2 := 0;
   END_IF;
   IF #in21 THEN
       #out2 := 1;
   END_IF;
   IF #in22 THEN
       #out2 := 2;
   END_IF;
   IF #in23 THEN
       #out2 := 3;
   END_IF;
   IF #in24 THEN
       #out2 := 4;
   END_IF;
   IF #in25 THEN
       #out2 := 5;
   END_IF;
END_FUNCTION

FUNCTION "input_timers" : Void   // FC2, SCL
{ S7_Optimized_Access := 'TRUE' }